// TIA Portal project "Pozycjoner_v7" (V15.1)

(* hardware
DEVICE "PLC"  S7-1200 Station
   slot 0: "Rack_0"  S7-1200 Rack  Rack  V1.0
   slot 1: "PLC"  CPU 1212C AC/DC/Rly  6ES7 212-1BE40-0XB0  V4.3
   slot 2: "DIO"  6ES7 223-1BH32-0XB0  V2.0
DEVICE "HMI"  KTP700 Basic PN
   slot 0: "HMI"  KTP700 Basic PN  6AV2 123-2GB03-0AX0  15.1.0.0
   slot 1: "HMI_RT"  KTP700 Basic PN  6AV2 123-2GB03-0AX0  15.1.0.0
   slot 5: "HMI.IE_CP_1"  PROFINET Interface  15.0.1.0
      slot 1: "PROFINET Interface_1"  PROFINET Interface
         slot 1: "Port_1"  Port
DEVICE "Axis_Y"  GSD.Device.PN
   slot 0: "Rack"  Rack  V1.0
   slot 0: "Axis_Y"  SINAMICS V90 PN V1.0  6SL3 210-5Fxxx-xxFx  V1.00
      slot 0: "SINAMICS V90 PN V1.0"  SINAMICS V90 PN V1.0
      slot 1: "PN-IO"  PN-IO
         slot 1: "Port 1"  Port 1
         slot 2: "Port 2"  Port 2
      slot 1: "Drive"  Drive
         slot 0: "Module Access Point"  Module Access Point
         slot 1: "without PROFIsafe"  without PROFIsafe
   slot 2: "SIEMENS telegram 111, PZD-12/12"  SIEMENS telegram 111, PZD-12/12
DEVICE "AXIS_X"  GSD.Device.PN
   slot 0: "Rack"  Rack  V1.0
   slot 0: "Axis_X"  SINAMICS V90 PN V1.0  6SL3 210-5Fxxx-xxFx  V1.00
      slot 0: "SINAMICS V90 PN V1.0"  SINAMICS V90 PN V1.0
      slot 1: "PN-IO"  PN-IO
         slot 1: "Port 1"  Port 1
         slot 2: "Port 2"  Port 2
      slot 1: "Drive"  Drive
         slot 0: "Module Access Point"  Module Access Point
         slot 1: "without PROFIsafe"  without PROFIsafe
   slot 2: "SIEMENS telegram 111, PZD-12/12"  SIEMENS telegram 111, PZD-12/12
DEVICE "Axis_Z"  GSD.Device.PN
   slot 0: "Rack"  Rack  V1.0
   slot 0: "Axis_Z"  SINAMICS V90 PN V1.0  6SL3 210-5Fxxx-xxFx  V1.00
      slot 0: "SINAMICS V90 PN V1.0"  SINAMICS V90 PN V1.0
      slot 1: "PN-IO"  PN-IO
         slot 1: "Port 1"  Port 1
         slot 2: "Port 2"  Port 2
      slot 1: "Drive"  Drive
         slot 0: "Module Access Point"  Module Access Point
         slot 1: "without PROFIsafe"  without PROFIsafe
   slot 2: "SIEMENS telegram 111, PZD-12/12"  SIEMENS telegram 111, PZD-12/12
*)

// ===== PLC "PLC"  CPU 1212C AC/DC/Rly =====
// protected blocks, not shown: "FB_Axis", "FB_DriveParameterCheck", "FB_SinaPara_S", "FB_SinaPos"

VAR_GLOBAL   // PLC tag table "Default tag table"
   "System_Byte" AT %MB0 : Byte;
   "FirstScan" AT %M0.0 : Bool;
   "DiagStatusUpdate" AT %M0.1 : Bool;
   "AlwaysTRUE" AT %M0.2 : Bool;
   "AlwaysFALSE" AT %M0.3 : Bool;
   "Clock_Byte" AT %MB1 : Byte;
   "Clock_10Hz" AT %M1.0 : Bool;
   "Clock_5Hz" AT %M1.1 : Bool;
   "Clock_2.5Hz" AT %M1.2 : Bool;
   "Clock_2Hz" AT %M1.3 : Bool;
   "Clock_1.25Hz" AT %M1.4 : Bool;
   "Clock_1Hz" AT %M1.5 : Bool;
   "Clock_0.625Hz" AT %M1.6 : Bool;
   "Clock_0.5Hz" AT %M1.7 : Bool;
   "Tag_1" AT %Q0.0 : Bool;
   "Laser Sensor" AT %I0.0 : Bool;
END_VAR

VAR_GLOBAL   // PLC tag table "IO"
   "Inductive_Sensor_4" AT %I8.0 : Bool;
   "Inductive_Sensor_3" AT %I8.1 : Bool;
   "Inductive_Sensor_2" AT %I8.2 : Bool;
   "Inductive_Sensor_1" AT %I8.3 : Bool;
   "I8.4" AT %I8.4 : Bool;
   "Laser_Sensor" AT %I8.5 : Bool;
   "EStop_Fdb" AT %I8.6 : Bool;
   "I8.7" AT %I8.7 : Bool;
   "Electromagnet" AT %Q8.0 : Bool;
   "Q8.1" AT %Q8.1 : Bool;
   "Q8.2" AT %Q8.2 : Bool;
   "Q8.3" AT %Q8.3 : Bool;
   "Q8.4" AT %Q8.4 : Bool;
   "Q8.5" AT %Q8.5 : Bool;
   "Q8.6" AT %Q8.6 : Bool;
   "Q8.7" AT %Q8.7 : Bool;
   "Axis_X_ActualTorque" AT %IW114 : Int;
   "Axis_Y_ActualTorque" AT %IW90 : Int;
   "Axis_Z_ActualTorque" AT %IW138 : Int;
END_VAR

TYPE "UDT_SinaPos"
   STRUCT
      ModePos : Int := 0;   // Settings of the mode
      EnableAxis : Bool := 0;   // 1 = Enable the drive
      CancelTraversing : Bool := 1;   // 0 = Reject active traverse task
      IntermediateStop : Bool := 1;   // 0 = Intermediate STOP of traverse command
      Positive : Bool := 0;   // 1 = Direction positive
      Negative : Bool := 0;   // 1 = Direction negative
      Jog1 : Bool := 0;   // 1 = Use jog 1 (direction / speed)
      Jog2 : Bool := 0;   // 1 = Use jog 2 (direction / speed)
      FlyRef : Bool := 0;   // 1 = Start flying reference function
      AckError : Bool := 0;   // 1 = Acknowledge of errors
      ExecuteMode : Bool := 0;   // 0-->1 = Start the mode
      Position : DInt := 0;   // Position of the MDI mode or setting of traversing block
      Velocity : DInt := 0;   // MDI velocity
      OverV : Int := 100;   // Override of velocity in [%] --> 4000h=100%
      OverAcc : Int := 100;   // Override of acceleration in [%] --> 4000h=100%
      OverDec : Int := 100;   // Override of deceleration in [%] --> 4000h=100%
      ConfigEPos : DWord := 16#0000_0003;   // binary programmed input to control all functions in the telegram without its own function block input
      HWIDSTW : Hw_Io := 0;   // Hardware Identifer set point slot
      HWIDZSW : Hw_Io := 0;   // Hardware Identifer actual value slot
      AxisEnabled : Bool := 0;   // 1= Axis in operation
      AxisPosOk : Bool := 0;   // 1= Position setpoint reached
      AxisSpFixed : Bool := false;   // 1= Setpoint fixed (Attention: Dependence on SINAMICS firmware)
      AxisRef : Bool := 0;   // 1= Reference point set
      AxisWarn : Bool := 0;   // 1= Axis alarm / warning present
      AxisError : Bool := 0;   // 1= Axis fault present
      Lockout : Bool := 0;   // 1= Axis in lockout state
      ActVelocity : DInt := 0;   // Actual drive speed (has to be normed with p2000 --> 40000000h = 100%)
      ActPosition : DInt := 0;   // Actual position in [LU]
      ActMode : Int := 0;   // Active EPos mode
      EPosZSW1 : Word := 0;   // Status of EPOS ZSW1
      EPosZSW2 : Word := 0;   // Status of EPOS ZSW2
      ActWarn : Word := 0;   // Actual number of warning
      ActFault : Word := 0;   // Actual number of error
      Error : Bool := 0;   // 1 = Error (FB and Infeed)
      Status : Word := 0;   // Status output (7002 = FB in operation; 8xxx = error description - read the manual)
      DiagID : Word := 0;   // Error codes of the cyclic system funtion blocks DPWR / DPRD_DAT
   END_STRUCT;
END_TYPE

TYPE "UDT_AxisConfiguration"
   STRUCT
      Siemens_Telegram : Hw_Io;   // Siemens Telegram Hardware Identifier
      DriveModule_AccessPoint : Hw_Io;   // Drive Module Access Point Hardware Identifier
      VelocityLimitCW : Real;   // CW Velocity limit
      VelocityLimitCCW : Real;   // CCW Velocity limit
      MaxVelocity : Real;   // Max Velocity limit
      TorqueLimit : Real;   // TorqueLimit
      SoftLimitSwitchCW : DInt;   // Software limit switch CW
      SoftLimitSwitchCCW : DInt;   // Software limit switch CCW
      RefTorquePos : Real;   // Referencing Torque Positive Direction
      RefTorqueNeg : Real;   // Referencing Torque Negative Direction
   END_STRUCT;
END_TYPE

TYPE "UDT_AxisStatus"
   STRUCT
      Enabled : Bool;   // Axis Enabled
      PositionSetpoint : DInt;   // Target Position (LU)
      VelocitySetpoint : DInt;   // Commanded Postion (LU/s)
      PositionReached : Bool;   // Position Reached Indication
      Referenced : Bool;   // Axis Referenced
      ActualVelocity : Real;   // Actual Velocity (mm/s)
      ActualPosition : Real;   // Actual Position (mm)
      LimitCW : Real;   // Limit Position Clockwise Direction (mm)
      LimitCCW : Real;   // Limit Position Counterclockwise Direction (mm)
      Error : Bool;   // Error Present
      ParamCheckError : Bool;   // Error Parameter Check
      Warning : Bool;   // Warning Present
      ErrorCode : Word;   // Error Code
      WarningCode : Word;   // Warning Code
      InvalidPosition : Bool;   // Invalid Commanded Position
      InvalidVelocity : Bool;   // Invalid Commanded Velocity
   END_STRUCT;
END_TYPE

TYPE "UDT_AxisControl"
   STRUCT
      JogActivate : Bool;   // Activate Jog Movement
      JogCW : Bool;   // Jog in Clockwise Direction
      JogCCW : Bool;   // Jog in Counterclockwise Direction
      SetReference : Bool;   // Start Axis Referencing
      ReqPosition : Real;   // Requested Position (mm)
      ReqVelocity : Real;   // Requested Velocity (mm/s)
      Start : Bool;   // Start Movement Command
      Stop : Bool;   // Stop Active Movement
   END_STRUCT;
END_TYPE

// folder: Displacement/Average Position

DATA_BLOCK "DB_AdditionalValues"   // DB16
{ S7_Optimized_Access := 'TRUE' }
VERSION : 0.1
// stored: InstanceOfName FB_AdditionalValues
"FB_AdditionalValues"
BEGIN
END_DATA_BLOCK

DATA_BLOCK "DB_Average positions"   // DB57
{ S7_Optimized_Access := 'TRUE' }
VERSION : 0.1
// stored: InstanceOfName FB_Average positions
"FB_Average positions"
BEGIN
END_DATA_BLOCK

// folder: Displacement/Center Point Calculation

DATA_BLOCK "DB_Falling_Edge"   // DB17
{ S7_Optimized_Access := 'TRUE' }
VERSION : 0.1
// stored: InstanceOfName FB_Falling_Edge
"FB_Falling_Edge"
BEGIN
END_DATA_BLOCK

// folder: Displacement/Center Point Calculation/Line2

DATA_BLOCK "DB_Line2"   // DB19
{ S7_Optimized_Access := 'TRUE' }
VERSION : 0.1
// stored: InstanceOfName FB_Line2
"FB_Line2"
BEGIN
END_DATA_BLOCK

// folder: Displacement/Center Point Calculation/Line3

DATA_BLOCK "DB_Line3"   // DB53
{ S7_Optimized_Access := 'TRUE' }
VERSION : 0.1
// stored: InstanceOfName FB_Line3
"FB_Line3"
BEGIN
END_DATA_BLOCK

// folder: Displacement/Object displacement

DATA_BLOCK "DB_Displacement"   // DB46
{ S7_Optimized_Access := 'TRUE' }
VERSION : 0.1
// stored: InstanceOfName FB_Displacement
"FB_Displacement"
BEGIN
END_DATA_BLOCK

// folder: Displacement/Object displacement/Inductive Sensors

DATA_BLOCK "DB_Inductive_Sensors"   // DB38
{ S7_Optimized_Access := 'TRUE' }
VERSION : 0.1
// stored: InstanceOfName FB_Inductive_Sensors
"FB_Inductive_Sensors"
BEGIN
END_DATA_BLOCK

// folder: Displacement/Object displacement/Velocity

DATA_BLOCK "DB_Velocity"   // DB40
{ S7_Optimized_Access := 'TRUE' }
VERSION : 0.1
// stored: InstanceOfName Velocity
"Velocity"
BEGIN
END_DATA_BLOCK

// folder: Drivers Parameters

DATA_BLOCK "DB_Interrupts"   // DB13
{ S7_Optimized_Access := 'TRUE' }
VERSION : 0.1
   VAR
      REInterrupt : Bool;   // Set when rising edge was detected
      FEInterrupt : Bool;   // Set when falling edge was detected
      GeneralCounter : Int;   // It shows which part of the program is performing
      RECounter : Int;
      FECounter : Int;   // The First Falling Edge Counter
      CountDown2 : Int;   // The Second Falling Edge Counter
      X2_positions : Array[0..10] of Real;   // X positions of the first falling edge
      Y2_positions : Array[0..10] of Real;   // Y positions of the first falling edge
      X4_positions : Array[0..20] of Real;   // X positions of the second falling edge
      Y4_positions : Array[0..20] of Real;   // Y positions of the second falling edge
      Positions : Struct
         "1" : Struct
            X : Real;
            Y : Real;
         END_STRUCT;
         "2" : Struct
            X : Real;
            Y : Real;
         END_STRUCT;
         "3" : Struct
            X : Real;
            Y : Real;
         END_STRUCT;
         "4" : Struct
            X : Real;
            Y : Real;
         END_STRUCT;
         "4*" : Struct
            X : Real;
            Y : Real;
         END_STRUCT;
         "5" : Struct
            X : Real;
            Y : Real;
         END_STRUCT;
         "6" : Struct
            X : Real;
            Y : Real;
         END_STRUCT;
         "4**" : Struct
            X : Real;
            Y : Real;
         END_STRUCT;
      END_STRUCT;
   END_VAR
BEGIN
END_DATA_BLOCK

DATA_BLOCK "DB_Drivers"   // DB14
{ S7_Optimized_Access := 'TRUE' }
VERSION : 0.1
// stored: InstanceOfName FB_Drivers
"FB_Drivers"
BEGIN
END_DATA_BLOCK

DATA_BLOCK "DB_Drivers_Interrupt"   // DB36
{ S7_Optimized_Access := 'TRUE' }
VERSION : 0.1
// stored: InstanceOfName FB_Drivers_Interrupt
"FB_Drivers_Interrupt"
BEGIN
END_DATA_BLOCK

// folder: Error

DATA_BLOCK "DB_Error"   // DB30
{ S7_Optimized_Access := 'TRUE' }
VERSION : 0.1
// stored: InstanceOfName FB_Error
"FB_Error"
BEGIN
END_DATA_BLOCK

// folder: HMI

DATA_BLOCK "DB_HMI"   // DB3
{ S7_Optimized_Access := 'TRUE' }
VERSION : 0.1
   VAR
      Reset : Bool;
      Searching : Bool;
      Enable : Bool;
      StartPosition : Bool;
      Interrupt : Bool;
      Electromagnet : Bool;
      AxisStatus : Array[0..2] of "UDT_AxisStatus";
      AxisControl : Array[0..2] of "UDT_AxisControl";
      MidPosCounting : Bool;
      AvailablePlace : Int;
      Error : Bool;
      "Start/Enable" : Bool;
      ItemwasFound : Bool;
      GrabbingTheItem : Bool;
      StartPositionReached : Bool;
      MovingToStartPosition : Bool;
      ErrorState : Int;
      ResetError : Bool;
      ErrorHMI : Bool;
      ResetSpace : Bool;
      PlaceOcc : Struct
         S1 : Bool;
         S2 : Bool;
         S3 : Bool;
         S4 : Bool;
      END_STRUCT;
      Returning : Bool;
      InvalidPosition : Bool;
      InvalidItem : Bool;
   END_VAR
BEGIN
   // AxisStatus[0] : X Axis
   // AxisStatus[1] : Y Axis
   // AxisStatus[2] : Z Axis
END_DATA_BLOCK

// folder: Instances

DATA_BLOCK "DB_Configuration"   // DB2
{ S7_Optimized_Access := 'TRUE' }
VERSION : 0.1
   VAR
      Axis_X : "UDT_AxisConfiguration";
      Axis_Y : "UDT_AxisConfiguration";
      Axis_Z : "UDT_AxisConfiguration";
   END_VAR
BEGIN
   Axis_X.Siemens_Telegram := 302;
   Axis_X.VelocityLimitCW := 400.0;
   Axis_X.TorqueLimit := 3.822;
   Axis_X.SoftLimitSwitchCW := 0;
   Axis_X.SoftLimitSwitchCCW := 0;
   Axis_X.VelocityLimitCCW := -400.0;
   Axis_X.MaxVelocity := 450.0;
   Axis_Y.VelocityLimitCW := 300.0;
   Axis_Y.VelocityLimitCCW := -300.0;
   Axis_Y.MaxVelocity := 350.0;
   Axis_Y.TorqueLimit := 3.822;
   Axis_Y.SoftLimitSwitchCW := 0;
   Axis_Y.SoftLimitSwitchCCW := 0;
   Axis_Y.Siemens_Telegram := 301;
   Axis_Z.Siemens_Telegram := 303;
   Axis_Z.VelocityLimitCW := 40.0;
   Axis_Z.VelocityLimitCCW := -40.0;
   Axis_Z.MaxVelocity := 60.0;
   Axis_Z.TorqueLimit := 0.504;
   Axis_Z.SoftLimitSwitchCW := 0;
   Axis_Z.SoftLimitSwitchCCW := 0;
   Axis_X.RefTorquePos := 0.4;
   Axis_X.RefTorqueNeg := -0.4;
   Axis_Y.RefTorquePos := 1.0;
   Axis_Y.RefTorqueNeg := -1.0;
   Axis_Z.RefTorquePos := 0.03;
   Axis_Z.RefTorqueNeg := -0.03;
   Axis_X.DriveModule_AccessPoint := 288;
   Axis_Y.DriveModule_AccessPoint := 279;
   Axis_Z.DriveModule_AccessPoint := 298;
END_DATA_BLOCK

// folder: RESET

DATA_BLOCK "DB_RESET"   // DB15
{ S7_Optimized_Access := 'TRUE' }
VERSION : 0.1
// stored: InstanceOfName FB_RESET
"FB_RESET"
BEGIN
END_DATA_BLOCK

// folder: Searching Mode

DATA_BLOCK "DB_Searching"   // DB5
{ S7_Optimized_Access := 'TRUE' }
VERSION : 0.1
// stored: InstanceOfName FB_Searching
"FB_Searching"
BEGIN
END_DATA_BLOCK

// folder: Searching Mode/Movement

DATA_BLOCK "DB_Movement"   // DB12
{ S7_Optimized_Access := 'TRUE' }
VERSION : 0.1
// stored: InstanceOfName FB_Movement
"FB_Movement"
BEGIN
END_DATA_BLOCK

// folder: Searching Mode/Starting Position

DATA_BLOCK "DB_StartingPosition"   // DB8
{ S7_Optimized_Access := 'TRUE' }
VERSION : 0.1
// stored: InstanceOfName FB_Starting Position
"FB_Starting Position"
BEGIN
END_DATA_BLOCK

// folder: System blocks/Program resources

DATA_BLOCK "IEC_Timer_0_DB_1"   // DB9
{ S7_Optimized_Access := 'TRUE' }
AUTHOR : Simatic
FAMILY : IEC
NAME : IEC_TMR
VERSION : 1.0
// stored: InstanceOfName IEC_TIMER
"IEC_TIMER"
BEGIN
END_DATA_BLOCK

DATA_BLOCK "IEC_Timer_0_DB_2"   // DB10
{ S7_Optimized_Access := 'TRUE' }
AUTHOR : Simatic
FAMILY : IEC
NAME : IEC_TMR
VERSION : 1.0
// stored: InstanceOfName IEC_TIMER
"IEC_TIMER"
BEGIN
END_DATA_BLOCK

DATA_BLOCK "IEC_Timer_0_DB_3"   // DB11
{ S7_Optimized_Access := 'TRUE' }
AUTHOR : Simatic
FAMILY : IEC
NAME : IEC_TMR
VERSION : 1.0
// stored: InstanceOfName IEC_TIMER
"IEC_TIMER"
BEGIN
END_DATA_BLOCK

DATA_BLOCK "IEC_Timer_0_DB_5"   // DB18
{ S7_Optimized_Access := 'TRUE' }
AUTHOR : Simatic
FAMILY : IEC
NAME : IEC_TMR
VERSION : 1.0
// stored: InstanceOfName IEC_TIMER
"IEC_TIMER"
BEGIN
END_DATA_BLOCK

DATA_BLOCK "IEC_Timer_0_DB_19"   // DB20
{ S7_Optimized_Access := 'TRUE' }
AUTHOR : Simatic
FAMILY : IEC
NAME : IEC_TMR
VERSION : 1.0
// stored: InstanceOfName IEC_TIMER
"IEC_TIMER"
BEGIN
END_DATA_BLOCK

DATA_BLOCK "IEC_Timer_0_DB_6"   // DB21
{ S7_Optimized_Access := 'TRUE' }
AUTHOR : Simatic
FAMILY : IEC
NAME : IEC_TMR
VERSION : 1.0
// stored: InstanceOfName IEC_TIMER
"IEC_TIMER"
BEGIN
END_DATA_BLOCK

DATA_BLOCK "IEC_Timer_0_DB_4"   // DB22
{ S7_Optimized_Access := 'TRUE' }
AUTHOR : Simatic
FAMILY : IEC
NAME : IEC_TMR
VERSION : 1.0
// stored: InstanceOfName IEC_TIMER
"IEC_TIMER"
BEGIN
END_DATA_BLOCK

DATA_BLOCK "IEC_Timer_0_DB_7"   // DB23
{ S7_Optimized_Access := 'TRUE' }
AUTHOR : Simatic
FAMILY : IEC
NAME : IEC_TMR
VERSION : 1.0
// stored: InstanceOfName IEC_TIMER
"IEC_TIMER"
BEGIN
END_DATA_BLOCK

DATA_BLOCK "IEC_Timer_0_DB_8"   // DB24
{ S7_Optimized_Access := 'TRUE' }
AUTHOR : Simatic
FAMILY : IEC
NAME : IEC_TMR
VERSION : 1.0
// stored: InstanceOfName IEC_TIMER
"IEC_TIMER"
BEGIN
END_DATA_BLOCK

DATA_BLOCK "IEC_Timer_0_DB_9"   // DB25
{ S7_Optimized_Access := 'TRUE' }
AUTHOR : Simatic
FAMILY : IEC
NAME : IEC_TMR
VERSION : 1.0
// stored: InstanceOfName IEC_TIMER
"IEC_TIMER"
BEGIN
END_DATA_BLOCK

DATA_BLOCK "IEC_Timer_0_DB_10"   // DB26
{ S7_Optimized_Access := 'TRUE' }
AUTHOR : Simatic
FAMILY : IEC
NAME : IEC_TMR
VERSION : 1.0
// stored: InstanceOfName IEC_TIMER
"IEC_TIMER"
BEGIN
END_DATA_BLOCK

DATA_BLOCK "IEC_Timer_0_DB_11"   // DB27
{ S7_Optimized_Access := 'TRUE' }
AUTHOR : Simatic
FAMILY : IEC
NAME : IEC_TMR
VERSION : 1.0
// stored: InstanceOfName IEC_TIMER
"IEC_TIMER"
BEGIN
END_DATA_BLOCK

DATA_BLOCK "IEC_Timer_0_DB_13"   // DB29
{ S7_Optimized_Access := 'TRUE' }
AUTHOR : Simatic
FAMILY : IEC
NAME : IEC_TMR
VERSION : 1.0
// stored: InstanceOfName IEC_TIMER
"IEC_TIMER"
BEGIN
END_DATA_BLOCK

DATA_BLOCK "IEC_Timer_0_DB_15"   // DB31
{ S7_Optimized_Access := 'TRUE' }
AUTHOR : Simatic
FAMILY : IEC
NAME : IEC_TMR
VERSION : 1.0
// stored: InstanceOfName IEC_TIMER
"IEC_TIMER"
BEGIN
END_DATA_BLOCK

DATA_BLOCK "IEC_Timer_0_DB_16"   // DB32
{ S7_Optimized_Access := 'TRUE' }
AUTHOR : Simatic
FAMILY : IEC
NAME : IEC_TMR
VERSION : 1.0
// stored: InstanceOfName IEC_TIMER
"IEC_TIMER"
BEGIN
END_DATA_BLOCK

DATA_BLOCK "IEC_Timer_0_DB_17"   // DB33
{ S7_Optimized_Access := 'TRUE' }
AUTHOR : Simatic
FAMILY : IEC
NAME : IEC_TMR
VERSION : 1.0
// stored: InstanceOfName IEC_TIMER
"IEC_TIMER"
BEGIN
END_DATA_BLOCK

DATA_BLOCK "IEC_Timer_0_DB_18"   // DB34
{ S7_Optimized_Access := 'TRUE' }
AUTHOR : Simatic
FAMILY : IEC
NAME : IEC_TMR
VERSION : 1.0
// stored: InstanceOfName IEC_TIMER
"IEC_TIMER"
BEGIN
END_DATA_BLOCK

DATA_BLOCK "IEC_Timer_0_DB_20"   // DB35
{ S7_Optimized_Access := 'TRUE' }
AUTHOR : Simatic
FAMILY : IEC
NAME : IEC_TMR
VERSION : 1.0
// stored: InstanceOfName IEC_TIMER
"IEC_TIMER"
BEGIN
END_DATA_BLOCK

DATA_BLOCK "IEC_Timer_0_DB_22"   // DB39
{ S7_Optimized_Access := 'TRUE' }
AUTHOR : Simatic
FAMILY : IEC
NAME : IEC_TMR
VERSION : 1.0
// stored: InstanceOfName IEC_TIMER
"IEC_TIMER"
BEGIN
END_DATA_BLOCK

DATA_BLOCK "IEC_Timer_0_DB_27"   // DB41
{ S7_Optimized_Access := 'TRUE' }
AUTHOR : Simatic
FAMILY : IEC
NAME : IEC_TMR
VERSION : 1.0
// stored: InstanceOfName IEC_TIMER
"IEC_TIMER"
BEGIN
END_DATA_BLOCK

DATA_BLOCK "IEC_Timer_0_DB_14"   // DB42
{ S7_Optimized_Access := 'TRUE' }
AUTHOR : Simatic
FAMILY : IEC
NAME : IEC_TMR
VERSION : 1.0
// stored: InstanceOfName IEC_TIMER
"IEC_TIMER"
BEGIN
END_DATA_BLOCK

DATA_BLOCK "IEC_Timer_0_DB_23"   // DB43
{ S7_Optimized_Access := 'TRUE' }
AUTHOR : Simatic
FAMILY : IEC
NAME : IEC_TMR
VERSION : 1.0
// stored: InstanceOfName IEC_TIMER
"IEC_TIMER"
BEGIN
END_DATA_BLOCK

DATA_BLOCK "IEC_Timer_0_DB_24"   // DB44
{ S7_Optimized_Access := 'TRUE' }
AUTHOR : Simatic
FAMILY : IEC
NAME : IEC_TMR
VERSION : 1.0
// stored: InstanceOfName IEC_TIMER
"IEC_TIMER"
BEGIN
END_DATA_BLOCK

DATA_BLOCK "IEC_Timer_0_DB_25"   // DB45
{ S7_Optimized_Access := 'TRUE' }
AUTHOR : Simatic
FAMILY : IEC
NAME : IEC_TMR
VERSION : 1.0
// stored: InstanceOfName IEC_TIMER
"IEC_TIMER"
BEGIN
END_DATA_BLOCK

DATA_BLOCK "IEC_Timer_0_DB_26"   // DB47
{ S7_Optimized_Access := 'TRUE' }
AUTHOR : Simatic
FAMILY : IEC
NAME : IEC_TMR
VERSION : 1.0
// stored: InstanceOfName IEC_TIMER
"IEC_TIMER"
BEGIN
END_DATA_BLOCK

DATA_BLOCK "IEC_Timer_0_DB_28"   // DB48
{ S7_Optimized_Access := 'TRUE' }
AUTHOR : Simatic
FAMILY : IEC
NAME : IEC_TMR
VERSION : 1.0
// stored: InstanceOfName IEC_TIMER
"IEC_TIMER"
BEGIN
END_DATA_BLOCK

DATA_BLOCK "IEC_Timer_0_DB_29"   // DB49
{ S7_Optimized_Access := 'TRUE' }
AUTHOR : Simatic
FAMILY : IEC
NAME : IEC_TMR
VERSION : 1.0
// stored: InstanceOfName IEC_TIMER
"IEC_TIMER"
BEGIN
END_DATA_BLOCK

DATA_BLOCK "IEC_Timer_0_DB_30"   // DB50
{ S7_Optimized_Access := 'TRUE' }
AUTHOR : Simatic
FAMILY : IEC
NAME : IEC_TMR
VERSION : 1.0
// stored: InstanceOfName IEC_TIMER
"IEC_TIMER"
BEGIN
END_DATA_BLOCK

DATA_BLOCK "IEC_Timer_0_DB_31"   // DB51
{ S7_Optimized_Access := 'TRUE' }
AUTHOR : Simatic
FAMILY : IEC
NAME : IEC_TMR
VERSION : 1.0
// stored: InstanceOfName IEC_TIMER
"IEC_TIMER"
BEGIN
END_DATA_BLOCK

DATA_BLOCK "IEC_Timer_0_DB_32"   // DB52
{ S7_Optimized_Access := 'TRUE' }
AUTHOR : Simatic
FAMILY : IEC
NAME : IEC_TMR
VERSION : 1.0
// stored: InstanceOfName IEC_TIMER
"IEC_TIMER"
BEGIN
END_DATA_BLOCK

DATA_BLOCK "IEC_Timer_0_DB_34"   // DB55
{ S7_Optimized_Access := 'TRUE' }
AUTHOR : Simatic
FAMILY : IEC
NAME : IEC_TMR
VERSION : 1.0
// stored: InstanceOfName IEC_TIMER
"IEC_TIMER"
BEGIN
END_DATA_BLOCK

DATA_BLOCK "IEC_Timer_0_DB_35"   // DB56
{ S7_Optimized_Access := 'TRUE' }
AUTHOR : Simatic
FAMILY : IEC
NAME : IEC_TMR
VERSION : 1.0
// stored: InstanceOfName IEC_TIMER
"IEC_TIMER"
BEGIN
END_DATA_BLOCK

DATA_BLOCK "IEC_Timer_0_DB_36"   // DB58
{ S7_Optimized_Access := 'TRUE' }
AUTHOR : Simatic
FAMILY : IEC
NAME : IEC_TMR
VERSION : 1.0
// stored: InstanceOfName IEC_TIMER
"IEC_TIMER"
BEGIN
END_DATA_BLOCK

DATA_BLOCK "IEC_Timer_0_DB_37"   // DB59
{ S7_Optimized_Access := 'TRUE' }
AUTHOR : Simatic
FAMILY : IEC
NAME : IEC_TMR
VERSION : 1.0
// stored: InstanceOfName IEC_TIMER
"IEC_TIMER"
BEGIN
END_DATA_BLOCK

DATA_BLOCK "IEC_Timer_0_DB_38"   // DB60
{ S7_Optimized_Access := 'TRUE' }
AUTHOR : Simatic
FAMILY : IEC
NAME : IEC_TMR
VERSION : 1.0
// stored: InstanceOfName IEC_TIMER
"IEC_TIMER"
BEGIN
END_DATA_BLOCK

DATA_BLOCK "IEC_Timer_0_DB_39"   // DB61
{ S7_Optimized_Access := 'TRUE' }
AUTHOR : Simatic
FAMILY : IEC
NAME : IEC_TMR
VERSION : 1.0
// stored: InstanceOfName IEC_TIMER
"IEC_TIMER"
BEGIN
END_DATA_BLOCK

DATA_BLOCK "IEC_Timer_0_DB_40"   // DB62
{ S7_Optimized_Access := 'TRUE' }
AUTHOR : Simatic
FAMILY : IEC
NAME : IEC_TMR
VERSION : 1.0
// stored: InstanceOfName IEC_TIMER
"IEC_TIMER"
BEGIN
END_DATA_BLOCK

// folder: Displacement/Average Position

FUNCTION_BLOCK "FB_Average positions"   // FB17, LAD
{ S7_Optimized_Access := 'TRUE' }
VERSION : 0.1
   VAR
      AveragePosition : Struct
         X : Real;
         Y : Real;
      END_STRUCT;
      APwithOffsets : Struct
         X : Real;
         Y : Real;
      END_STRUCT;
      Ranges : Struct
         Xavg : Struct
            Min : Real;
            Max : Real;
         END_STRUCT;
         Yavg : Struct
            Min : Real;
            Max : Real;
         END_STRUCT;
         NewXavg : Struct
            Min : Real;
            Max : Real;
         END_STRUCT;
         NewYavg : Struct
            Min : Real;
            Max : Real;
         END_STRUCT;
         DiffX : Struct
            Min : Real;
            Max : Real;
         END_STRUCT;
      END_STRUCT;
      Positions : Struct
         "1" : Struct
            X : Real;
            Y : Real;
         END_STRUCT;
         "2" : Struct
            X : Real;
            Y : Real;
         END_STRUCT;
         "3" : Struct
            X : Real;
            Y : Real;
         END_STRUCT;
         "4" : Struct
            X : Real;
            Y : Real;
         END_STRUCT;
         New4 : Struct
            X : Real;
            Y : Real;
         END_STRUCT;
      END_STRUCT;
      NewAvegagePosition : Bool;
      "PosX+2" : Real;
   END_VAR
   VAR CONSTANT
      OffsetX : Real := 5.0;
      OffsetY : Real := 8.0;
      OffsetZ : Real := 86.5;
      RangeCen : Real := 2.5;
   END_VAR
   VAR_TEMP   // added for the SCL form of the ladder/FBD networks
      _w1 : Bool;
   END_VAR
BEGIN

REGION Network 1: Save values
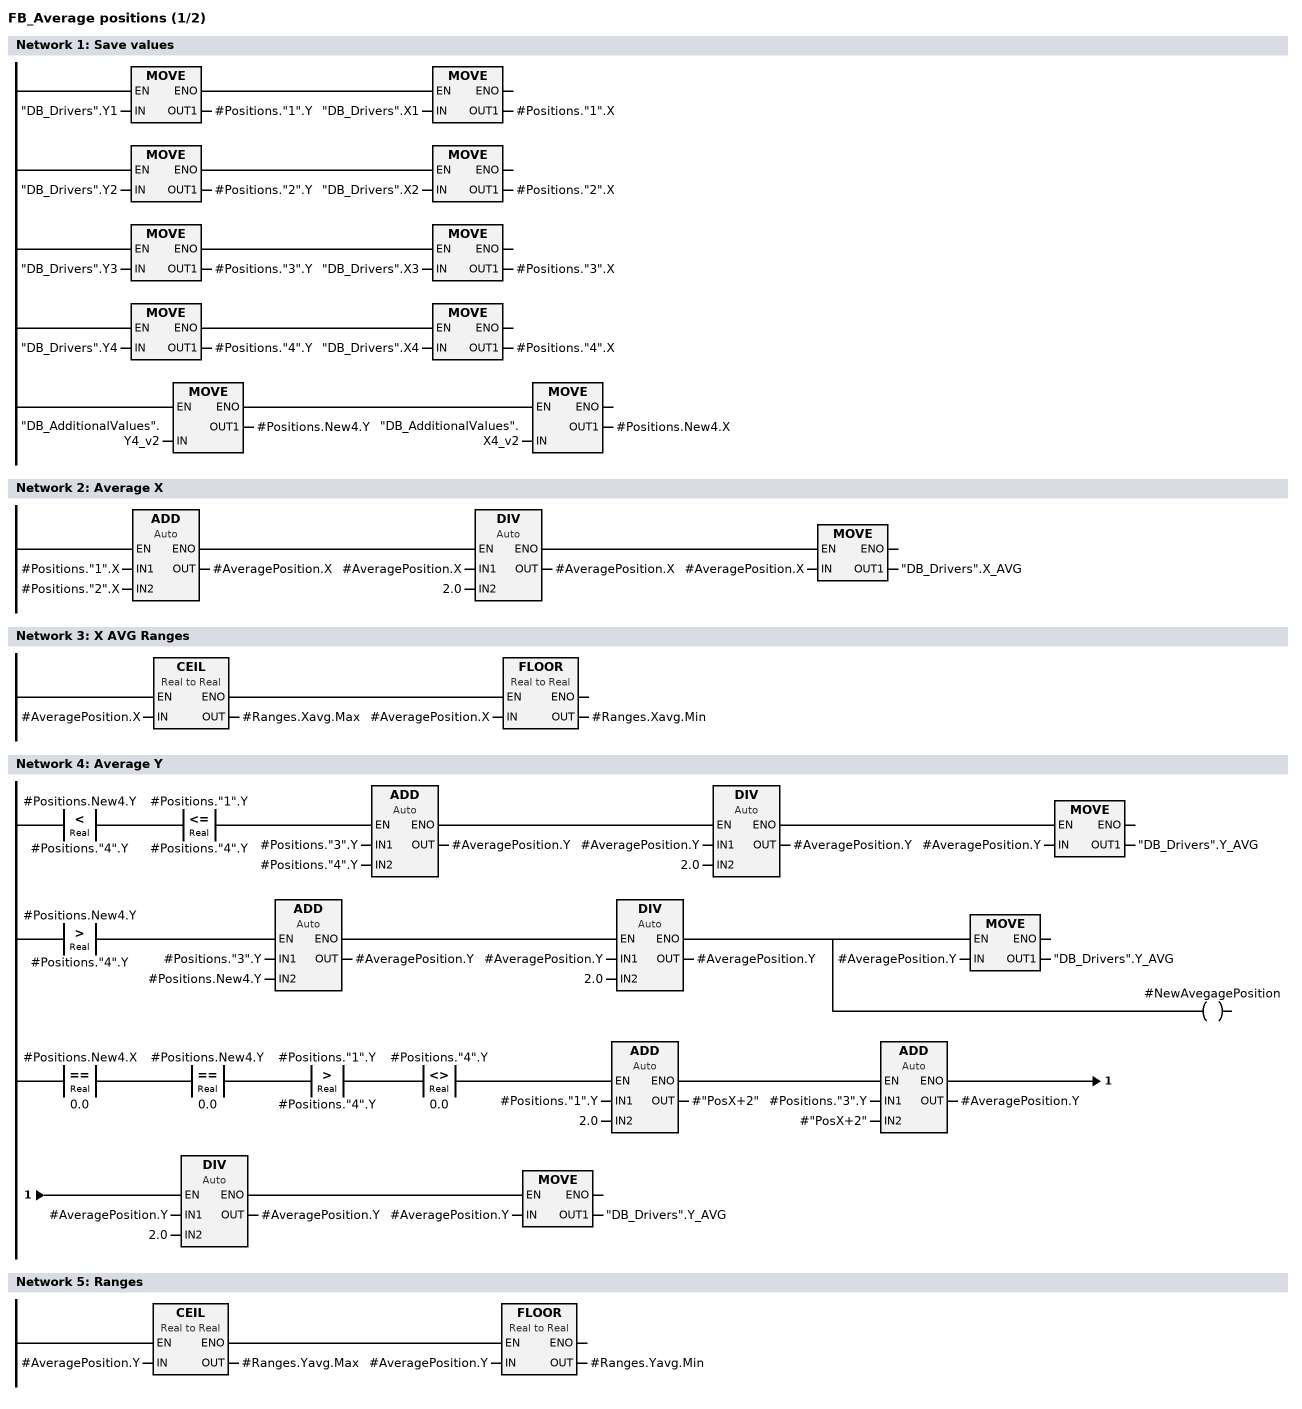
   RUNG wire#powerrail
      Move(in := "DB_Drivers".Y1, out1 => #Positions."1".Y)
      Move(in := "DB_Drivers".X1, out1 => #Positions."1".X)
   END_RUNG
   RUNG wire#powerrail
      Move(in := "DB_Drivers".Y2, out1 => #Positions."2".Y)
      Move(in := "DB_Drivers".X2, out1 => #Positions."2".X)
   END_RUNG
   RUNG wire#powerrail
      Move(in := "DB_Drivers".Y3, out1 => #Positions."3".Y)
      Move(in := "DB_Drivers".X3, out1 => #Positions."3".X)
   END_RUNG
   RUNG wire#powerrail
      Move(in := "DB_Drivers".Y4, out1 => #Positions."4".Y)
      Move(in := "DB_Drivers".X4, out1 => #Positions."4".X)
   END_RUNG
   RUNG wire#powerrail
      Move(in := "DB_AdditionalValues".Y4_v2, out1 => #Positions.New4.Y)
      Move(in := "DB_AdditionalValues".X4_v2, out1 => #Positions.New4.X)
   END_RUNG
   // the same network as SCL:
   #Positions."1".Y := "DB_Drivers".Y1;
   #Positions."1".X := "DB_Drivers".X1;
   #Positions."2".Y := "DB_Drivers".Y2;
   #Positions."2".X := "DB_Drivers".X2;
   #Positions."3".Y := "DB_Drivers".Y3;
   #Positions."3".X := "DB_Drivers".X3;
   #Positions."4".Y := "DB_Drivers".Y4;
   #Positions."4".X := "DB_Drivers".X4;
   #Positions.New4.Y := "DB_AdditionalValues".Y4_v2;
   #Positions.New4.X := "DB_AdditionalValues".X4_v2;
END_REGION

REGION Network 2: Average X
   RUNG wire#powerrail
      Add(in1 := #Positions."1".X, in2 := #Positions."2".X, out => #AveragePosition.X)
      Div(in1 := #AveragePosition.X, in2 := 2.0, out => #AveragePosition.X)
      Move(in := #AveragePosition.X, out1 => "DB_Drivers".X_AVG)
   END_RUNG
   // the same network as SCL:
   #AveragePosition.X := #Positions."1".X + #Positions."2".X;
   #AveragePosition.X := #AveragePosition.X / 2.0;
   "DB_Drivers".X_AVG := #AveragePosition.X;
END_REGION

REGION Network 3: X AVG Ranges
   #Ranges.Xavg.Max := CEIL(#AveragePosition.X);
   #Ranges.Xavg.Min := FLOOR(#AveragePosition.X);
END_REGION

REGION Network 4: Average Y
   RUNG wire#powerrail
      { S7_Templates := "SrcType := Real" } LT_Contact(in1 := #Positions.New4.Y, in2 := #Positions."4".Y)
      { S7_Templates := "SrcType := Real" } LE_Contact(in1 := #Positions."1".Y, in2 := #Positions."4".Y)
      Add(in1 := #Positions."3".Y, in2 := #Positions."4".Y, out => #AveragePosition.Y)
      Div(in1 := #AveragePosition.Y, in2 := 2.0, out => #AveragePosition.Y)
      Move(in := #AveragePosition.Y, out1 => "DB_Drivers".Y_AVG)
   END_RUNG
   RUNG wire#powerrail
      { S7_Templates := "SrcType := Real" } GT_Contact(in1 := #Positions.New4.Y, in2 := #Positions."4".Y)
      Add(in1 := #Positions."3".Y, in2 := #Positions.New4.Y, out => #AveragePosition.Y)
      Div(in1 := #AveragePosition.Y, in2 := 2.0, out => #AveragePosition.Y)
      wire#w1
      Move(in := #AveragePosition.Y, out1 => "DB_Drivers".Y_AVG)
   END_RUNG
   RUNG wire#w1
      Coil( #NewAvegagePosition )
   END_RUNG
   RUNG wire#powerrail
      { S7_Templates := "SrcType := Real" } EQ_Contact(in1 := #Positions.New4.X, in2 := 0.0)
      { S7_Templates := "SrcType := Real" } EQ_Contact(in1 := #Positions.New4.Y, in2 := 0.0)
      { S7_Templates := "SrcType := Real" } GT_Contact(in1 := #Positions."1".Y, in2 := #Positions."4".Y)
      { S7_Templates := "SrcType := Real" } NE_Contact(in1 := #Positions."4".Y, in2 := 0.0)
      Add(in1 := #Positions."1".Y, in2 := 2.0, out => #"PosX+2")
      Add(in1 := #Positions."3".Y, in2 := #"PosX+2", out => #AveragePosition.Y)
      Div(in1 := #AveragePosition.Y, in2 := 2.0, out => #AveragePosition.Y)
      Move(in := #AveragePosition.Y, out1 => "DB_Drivers".Y_AVG)
   END_RUNG
   // the same network as SCL:
   IF (#Positions.New4.Y < #Positions."4".Y) AND (#Positions."1".Y <= #Positions."4".Y) THEN
       #AveragePosition.Y := #Positions."3".Y + #Positions."4".Y;
       #AveragePosition.Y := #AveragePosition.Y / 2.0;
       "DB_Drivers".Y_AVG := #AveragePosition.Y;
   END_IF;
   #_w1 := #Positions.New4.Y > #Positions."4".Y;
   IF #_w1 THEN
       #AveragePosition.Y := #Positions."3".Y + #Positions.New4.Y;
       #AveragePosition.Y := #AveragePosition.Y / 2.0;
       "DB_Drivers".Y_AVG := #AveragePosition.Y;
   END_IF;
   #NewAvegagePosition := #_w1;
   IF (#Positions.New4.X = 0.0) AND (#Positions.New4.Y = 0.0) AND (#Positions."1".Y > #Positions."4".Y) AND (#Positions."4".Y <> 0.0) THEN
       #"PosX+2" := #Positions."1".Y + 2.0;
       #AveragePosition.Y := #Positions."3".Y + #"PosX+2";
       #AveragePosition.Y := #AveragePosition.Y / 2.0;
       "DB_Drivers".Y_AVG := #AveragePosition.Y;
   END_IF;
END_REGION

REGION Network 5: Ranges
   #Ranges.Yavg.Max := CEIL(#AveragePosition.Y);
   #Ranges.Yavg.Min := FLOOR(#AveragePosition.Y);
END_REGION

REGION Network 6: Ranges around center point
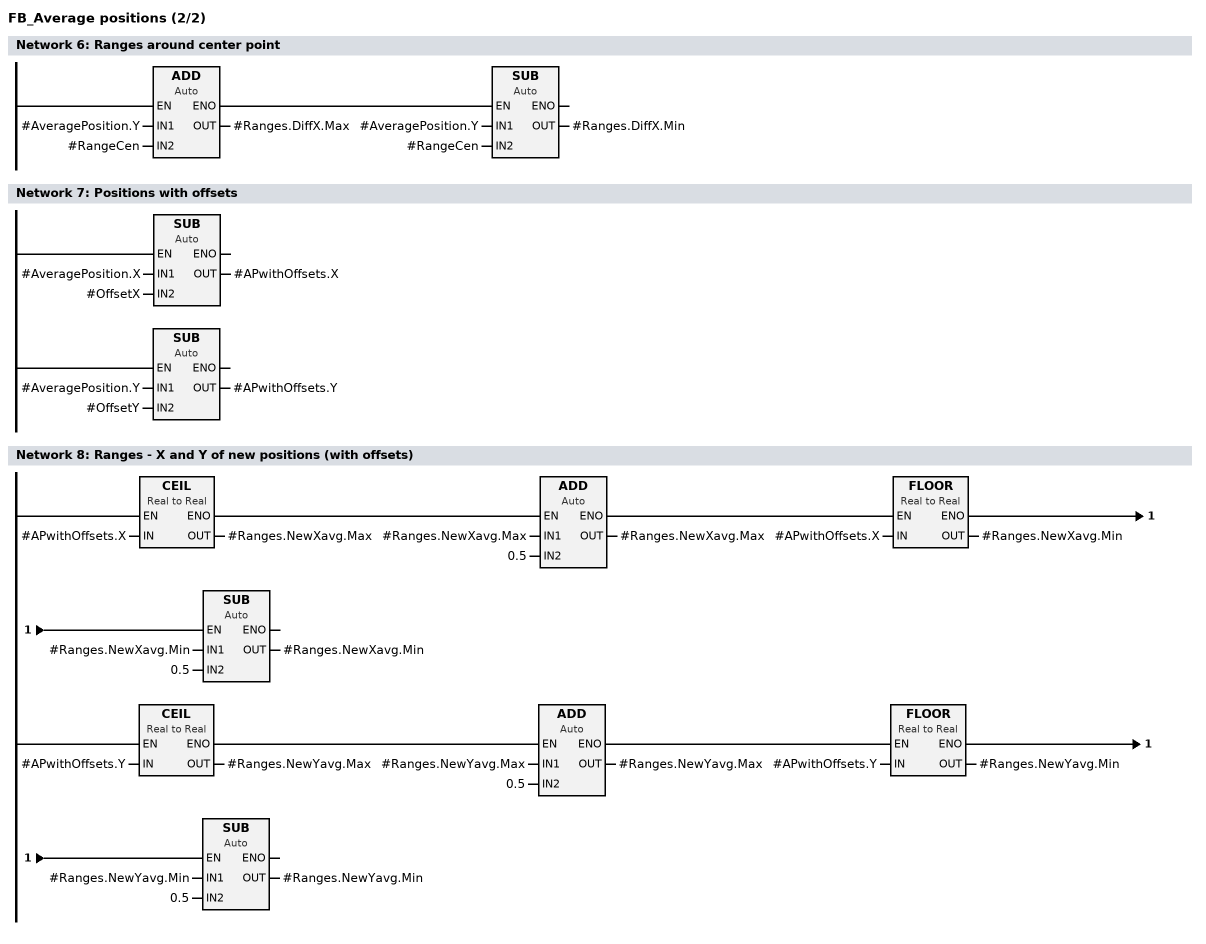
   RUNG wire#powerrail
      Add(in1 := #AveragePosition.Y, in2 := #RangeCen, out => #Ranges.DiffX.Max)
      Sub(in1 := #AveragePosition.Y, in2 := #RangeCen, out => #Ranges.DiffX.Min)
   END_RUNG
   // the same network as SCL:
   #Ranges.DiffX.Max := #AveragePosition.Y + #RangeCen;
   #Ranges.DiffX.Min := #AveragePosition.Y - #RangeCen;
END_REGION

REGION Network 7: Positions with offsets
   RUNG wire#powerrail
      Sub(in1 := #AveragePosition.X, in2 := #OffsetX, out => #APwithOffsets.X)
   END_RUNG
   RUNG wire#powerrail
      Sub(in1 := #AveragePosition.Y, in2 := #OffsetY, out => #APwithOffsets.Y)
   END_RUNG
   // the same network as SCL:
   #APwithOffsets.X := #AveragePosition.X - #OffsetX;
   #APwithOffsets.Y := #AveragePosition.Y - #OffsetY;
END_REGION

REGION Network 8: Ranges - X and Y of new positions (with offsets)
   #Ranges.NewXavg.Max := CEIL(#APwithOffsets.X);
   #Ranges.NewXavg.Max := #Ranges.NewXavg.Max + 0.5;
   #Ranges.NewXavg.Min := FLOOR(#APwithOffsets.X);
   #Ranges.NewXavg.Min := #Ranges.NewXavg.Min - 0.5;
   #Ranges.NewYavg.Max := CEIL(#APwithOffsets.Y);
   #Ranges.NewYavg.Max := #Ranges.NewYavg.Max + 0.5;
   #Ranges.NewYavg.Min := FLOOR(#APwithOffsets.Y);
   #Ranges.NewYavg.Min := #Ranges.NewYavg.Min - 0.5;
END_REGION
END_FUNCTION_BLOCK

// folder: Displacement/Center Point Calculation

FUNCTION_BLOCK "FB_AdditionalValues"   // FB8, LAD
{ S7_Optimized_Access := 'TRUE' }
VERSION : 0.1
   VAR
      UDT_AxisControl : Array[0..2] of "UDT_AxisControl";
      StopIncRE : Bool;   // Stop incremening
      DifX : Real;   // Difference between position X1 and X2
      SetPoint1Values : Bool;
      i : Int;
      "i-1" : Int;
      "i-2" : Int;
      "i+1" : Int;
      y1min : Int;
      y1max : Int;
      j : Int;
      "j-1" : Int;
      "j-2" : Int;
      "j+1" : Int;
      x3min : Int;
      x3max : Int;
      SetPoint3Values : Bool;
      X4_v2 : Real;
      Y4_v2 : Real;
      PtrigRE : Array[0..2] of Bool;
      StartFE : Array[0..5] of Bool;
      PtrigFE : Array[0..5] of Bool;
      Tim : Array[0..4] of Bool;
      Pulse : Array[0..1] of Bool;
   END_VAR
   VAR_TEMP   // added for the SCL form of the ladder/FBD networks
      _w1 : Bool;
      _w2 : Bool;
   END_VAR
BEGIN

REGION Network 1: Increment RisingEdge Counter
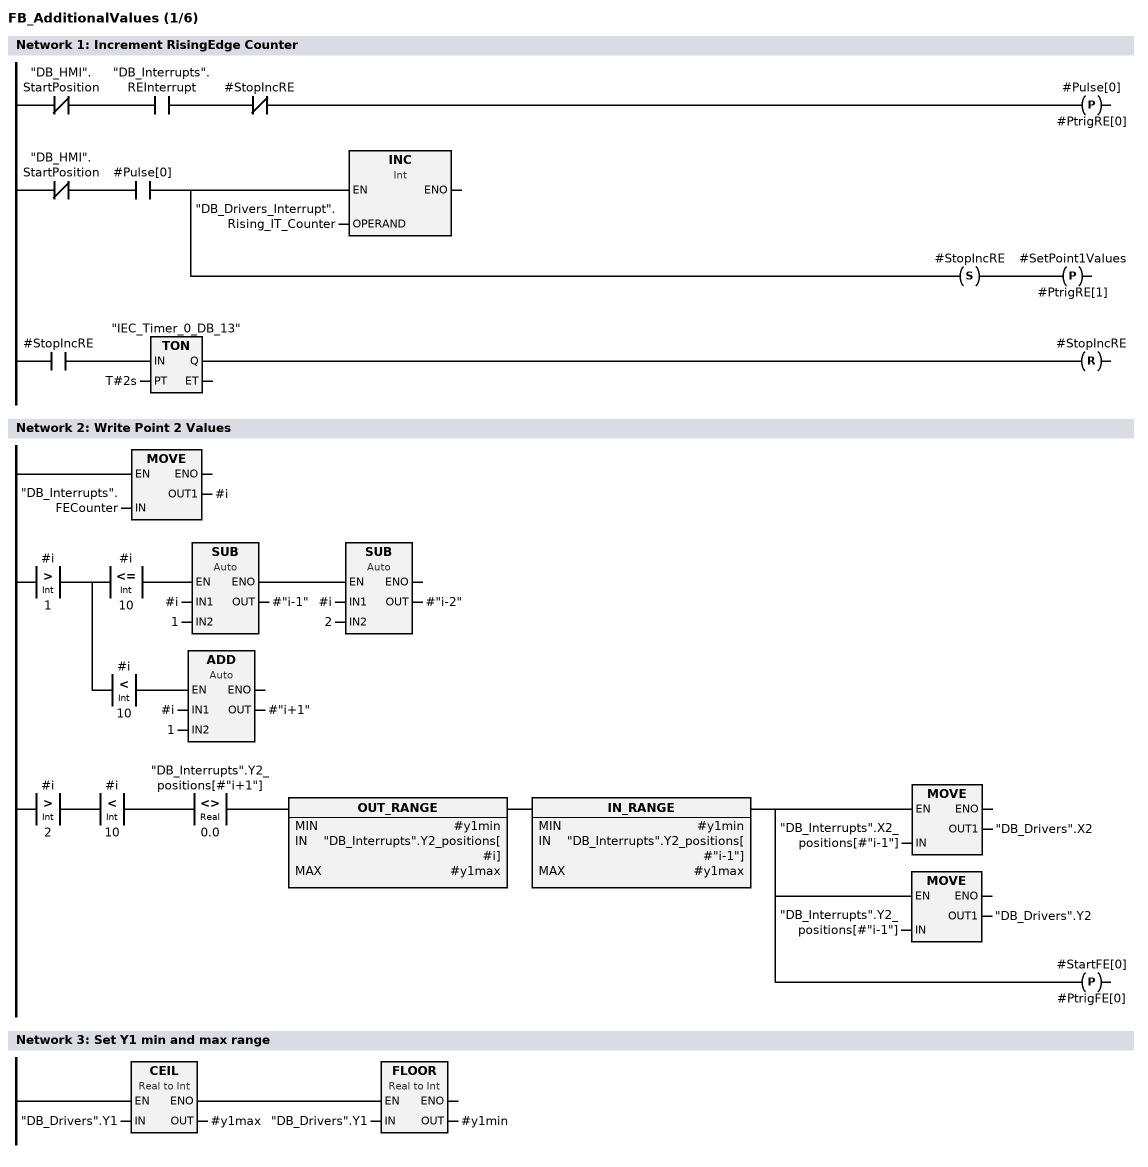
   #_w1 := NOT "DB_HMI".StartPosition AND "DB_Interrupts".REInterrupt AND NOT #StopIncRE;
   #Pulse[0] := #_w1 AND NOT #PtrigRE[0];   // rising edge
   #PtrigRE[0] := #_w1;
   #_w2 := NOT "DB_HMI".StartPosition AND #Pulse[0];
   IF #_w2 THEN
       "DB_Drivers_Interrupt".Rising_IT_Counter := "DB_Drivers_Interrupt".Rising_IT_Counter + 1;
       #StopIncRE := TRUE;
   END_IF;
   #SetPoint1Values := #_w2 AND NOT #PtrigRE[1];   // rising edge
   #PtrigRE[1] := #_w2;
   "IEC_Timer_0_DB_13".TON(IN := #StopIncRE, PT := T#2s);
   IF "IEC_Timer_0_DB_13".Q THEN #StopIncRE := FALSE; END_IF;
END_REGION

REGION Network 2: Write Point 2 Values
   #i := "DB_Interrupts".FECounter;
   #_w1 := #i > 1;
   IF #_w1 AND (#i <= 10) THEN
       #"i-1" := #i - 1;
       #"i-2" := #i - 2;
   END_IF;
   IF #_w1 AND (#i < 10) THEN #"i+1" := #i + 1; END_IF;
   #_w2 := (#i > 2) AND (#i < 10) AND ("DB_Interrupts".Y2_positions[#"i+1"] <> 0.0) AND (("DB_Interrupts".Y2_positions[#i] < #y1min) OR ("DB_Interrupts".Y2_positions[#i] > #y1max)) AND (#y1min <= "DB_Interrupts".Y2_positions[#"i-1"]) AND ("DB_Interrupts".Y2_positions[#"i-1"] <= #y1max);
   IF #_w2 THEN
       "DB_Drivers".X2 := "DB_Interrupts".X2_positions[#"i-1"];
       "DB_Drivers".Y2 := "DB_Interrupts".Y2_positions[#"i-1"];
   END_IF;
   #StartFE[0] := #_w2 AND NOT #PtrigFE[0];   // rising edge
   #PtrigFE[0] := #_w2;
END_REGION

REGION Network 3: Set Y1 min and max range
   #y1max := CEIL("DB_Drivers".Y1);
   #y1min := FLOOR("DB_Drivers".Y1);
END_REGION

REGION Network 4: Set Point 2 Values v2
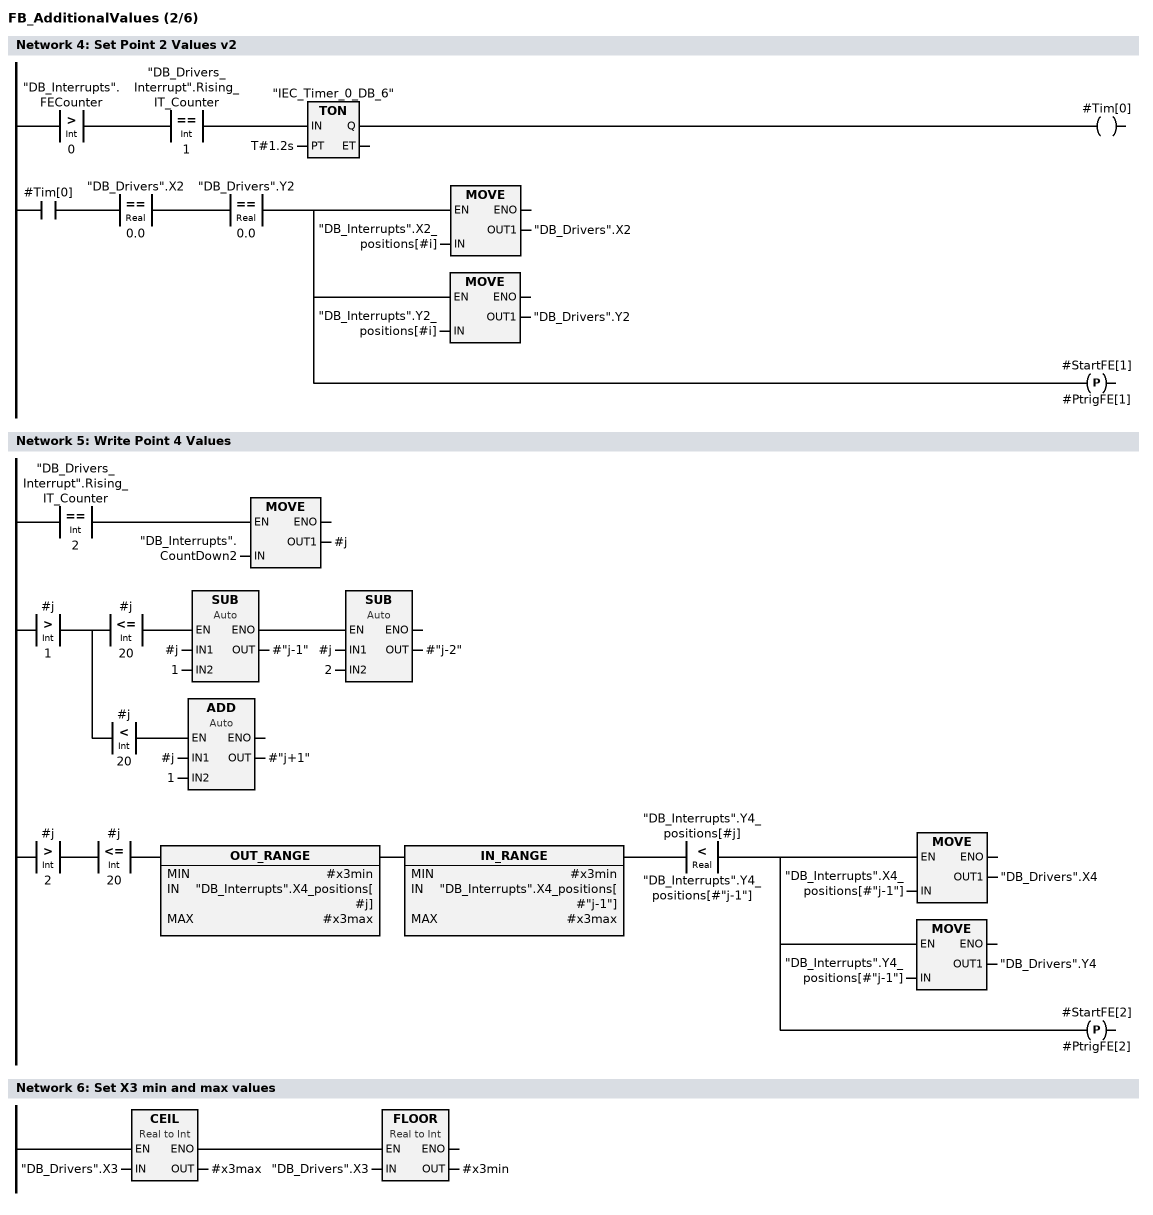
   "IEC_Timer_0_DB_6".TON(IN := ("DB_Interrupts".FECounter > 0) AND ("DB_Drivers_Interrupt".Rising_IT_Counter = 1),
                          PT := T#1.2s);
   #Tim[0] := "IEC_Timer_0_DB_6".Q;
   #_w1 := #Tim[0] AND ("DB_Drivers".X2 = 0.0) AND ("DB_Drivers".Y2 = 0.0);
   IF #_w1 THEN
       "DB_Drivers".X2 := "DB_Interrupts".X2_positions[#i];
       "DB_Drivers".Y2 := "DB_Interrupts".Y2_positions[#i];
   END_IF;
   #StartFE[1] := #_w1 AND NOT #PtrigFE[1];   // rising edge
   #PtrigFE[1] := #_w1;
END_REGION

REGION Network 5: Write Point 4 Values
   IF "DB_Drivers_Interrupt".Rising_IT_Counter = 2 THEN #j := "DB_Interrupts".CountDown2; END_IF;
   #_w1 := #j > 1;
   IF #_w1 AND (#j <= 20) THEN
       #"j-1" := #j - 1;
       #"j-2" := #j - 2;
   END_IF;
   IF #_w1 AND (#j < 20) THEN #"j+1" := #j + 1; END_IF;
   #_w2 := (#j > 2) AND (#j <= 20) AND (("DB_Interrupts".X4_positions[#j] < #x3min) OR ("DB_Interrupts".X4_positions[#j] > #x3max)) AND (#x3min <= "DB_Interrupts".X4_positions[#"j-1"]) AND ("DB_Interrupts".X4_positions[#"j-1"] <= #x3max) AND ("DB_Interrupts".Y4_positions[#j] < "DB_Interrupts".Y4_positions[#"j-1"]);
   IF #_w2 THEN
       "DB_Drivers".X4 := "DB_Interrupts".X4_positions[#"j-1"];
       "DB_Drivers".Y4 := "DB_Interrupts".Y4_positions[#"j-1"];
   END_IF;
   #StartFE[2] := #_w2 AND NOT #PtrigFE[2];   // rising edge
   #PtrigFE[2] := #_w2;
END_REGION

REGION Network 6: Set X3 min and max values
   #x3max := CEIL("DB_Drivers".X3);
   #x3min := FLOOR("DB_Drivers".X3);
END_REGION

REGION Network 7: Write Point 4 Values v2
   // Before it was 1s.